   "DB_SDC_EMS_TS_1_HMI_SEK[165].EMS[1]" : UDT_SDC_EMS_TS_STAT_HMI = PLC DB_SDC_EMS_TS_1_HMI.SEK[165].EMS[1] AT %DB3810.DBX29540.0, 1 s
   "DB_SDC_EMS_TS_1_HMI_SEK[166].EMS[1]" : UDT_SDC_EMS_TS_STAT_HMI = PLC DB_SDC_EMS_TS_1_HMI.SEK[166].EMS[1] AT %DB3810.DBX29720.0, 1 s
   "DB_SDC_EMS_TS_1_HMI_SEK[167].EMS[1]" : UDT_SDC_EMS_TS_STAT_HMI = PLC DB_SDC_EMS_TS_1_HMI.SEK[167].EMS[1] AT %DB3810.DBX29900.0, 1 s
   "DB_SDC_EMS_TS_1_HMI_SEK[168].EMS[1]" : UDT_SDC_EMS_TS_STAT_HMI = PLC DB_SDC_EMS_TS_1_HMI.SEK[168].EMS[1] AT %DB3810.DBX30080.0, 1 s
   "DB_SDC_EMS_TS_1_HMI_SEK[169].EMS[1]" : UDT_SDC_EMS_TS_STAT_HMI = PLC DB_SDC_EMS_TS_1_HMI.SEK[169].EMS[1] AT %DB3810.DBX30260.0, 1 s
   "DB_SDC_EMS_TS_1_HMI_SEK[170].EMS[1]" : UDT_SDC_EMS_TS_STAT_HMI = PLC DB_SDC_EMS_TS_1_HMI.SEK[170].EMS[1] AT %DB3810.DBX30440.0, 1 s
   "DB_SDC_EMS_TS_1_HMI_SEK[190].EMS[1]" : UDT_SDC_EMS_TS_STAT_HMI = PLC DB_SDC_EMS_TS_1_HMI.SEK[190].EMS[1] AT %DB3810.DBX34040.0, 1 s
   "DB_SDC_EMS_TS_1_HMI_SEK[191].EMS[1]" : UDT_SDC_EMS_TS_STAT_HMI = PLC DB_SDC_EMS_TS_1_HMI.SEK[191].EMS[1] AT %DB3810.DBX34220.0, 1 s
   "DB_SDC_EMS_TS_1_HMI_SEK[192].EMS[1]" : UDT_SDC_EMS_TS_STAT_HMI = PLC DB_SDC_EMS_TS_1_HMI.SEK[192].EMS[1] AT %DB3810.DBX34400.0, 1 s
   "DB_SDC_EMS_TS_1_HMI_SEK[193].EMS[1]" : UDT_SDC_EMS_TS_STAT_HMI = PLC DB_SDC_EMS_TS_1_HMI.SEK[193].EMS[1] AT %DB3810.DBX34580.0, 1 s
   "DB_SDC_EMS_TS_1_HMI_SEK[194].EMS[1]" : UDT_SDC_EMS_TS_STAT_HMI = PLC DB_SDC_EMS_TS_1_HMI.SEK[194].EMS[1] AT %DB3810.DBX34760.0, 1 s
   "DB_SDC_EMS_TS_1_HMI_SEK[195].EMS[1]" : UDT_SDC_EMS_TS_STAT_HMI = PLC DB_SDC_EMS_TS_1_HMI.SEK[195].EMS[1] AT %DB3810.DBX34940.0, 1 s
   "DB_SDC_EMS_TS_1_HMI_SEK[86].EMS[1]" : UDT_SDC_EMS_TS_STAT_HMI = PLC DB_SDC_EMS_TS_1_HMI.SEK[86].EMS[1] AT %DB3810.DBX15320.0, 1 s
   "DB_SDC_EMS_TS_1_HMI_SEK[87].EMS[1]" : UDT_SDC_EMS_TS_STAT_HMI = PLC DB_SDC_EMS_TS_1_HMI.SEK[87].EMS[1] AT %DB3810.DBX15500.0, 1 s
   "DB_SDC_EMS_TS_1_HMI_SEK[137].EMS[1]" : UDT_SDC_EMS_TS_STAT_HMI = PLC DB_SDC_EMS_TS_1_HMI.SEK[137].EMS[1] AT %DB3810.DBX24500.0, 1 s
   "DB_SDC_EMS_TS_1_HMI_SEK[136].EMS[1]" : UDT_SDC_EMS_TS_STAT_HMI = PLC DB_SDC_EMS_TS_1_HMI.SEK[136].EMS[1] AT %DB3810.DBX24320.0, 1 s
   "DB_SDC_EMS_TS_1_HMI_SEK[135].EMS[1]" : UDT_SDC_EMS_TS_STAT_HMI = PLC DB_SDC_EMS_TS_1_HMI.SEK[135].EMS[1] AT %DB3810.DBX24140.0, 1 s
   "DB_SDC_EMS_TS_1_HMI_SEK[134].EMS[1]" : UDT_SDC_EMS_TS_STAT_HMI = PLC DB_SDC_EMS_TS_1_HMI.SEK[134].EMS[1] AT %DB3810.DBX23960.0, 1 s

HMI tags "DB_SDC_EMS_TS_HMI_BA2"
   "DB_SDC_EMS_TS_1_HMI_SEK[99].EMS[1]" : UDT_SDC_EMS_TS_STAT_HMI = PLC DB_SDC_EMS_TS_1_HMI.SEK[99].EMS[1] AT %DB3810.DBX17660.0, 1 s
   "DB_SDC_EMS_TS_1_HMI_SEK[100].EMS[1](1)" : UDT_SDC_EMS_TS_STAT_HMI = PLC DB_SDC_EMS_TS_1_HMI.SEK[100].EMS[1] AT %DB3810.DBX17840.0, 1 s
   "DB_SDC_EMS_TS_1_HMI_SEK[101].EMS[1](1)" : UDT_SDC_EMS_TS_STAT_HMI = PLC DB_SDC_EMS_TS_1_HMI.SEK[101].EMS[1] AT %DB3810.DBX18020.0, 1 s
   "DB_SDC_EMS_TS_1_HMI_SEK[102].EMS[1](1)" : UDT_SDC_EMS_TS_STAT_HMI = PLC DB_SDC_EMS_TS_1_HMI.SEK[102].EMS[1] AT %DB3810.DBX18200.0, 1 s
   "DB_SDC_EMS_TS_1_HMI_SEK[103].EMS[1](1)" : UDT_SDC_EMS_TS_STAT_HMI = PLC DB_SDC_EMS_TS_1_HMI.SEK[103].EMS[1] AT %DB3810.DBX18380.0, 1 s
   "DB_SDC_EMS_TS_1_HMI_SEK[104].EMS[1](1)" : UDT_SDC_EMS_TS_STAT_HMI = PLC DB_SDC_EMS_TS_1_HMI.SEK[104].EMS[1] AT %DB3810.DBX18560.0, 1 s
   "DB_SDC_EMS_TS_1_HMI_SEK[105].EMS[1](1)" : UDT_SDC_EMS_TS_STAT_HMI = PLC DB_SDC_EMS_TS_1_HMI.SEK[105].EMS[1] AT %DB3810.DBX18740.0, 1 s
   "DB_SDC_EMS_TS_1_HMI_SEK[106].EMS[1](1)" : UDT_SDC_EMS_TS_STAT_HMI = PLC DB_SDC_EMS_TS_1_HMI.SEK[106].EMS[1] AT %DB3810.DBX18920.0, 1 s
   "DB_SDC_EMS_TS_1_HMI_SEK[107].EMS[1](1)" : UDT_SDC_EMS_TS_STAT_HMI = PLC DB_SDC_EMS_TS_1_HMI.SEK[107].EMS[1] AT %DB3810.DBX19100.0, 1 s
   "DB_SDC_EMS_TS_1_HMI_SEK[108].EMS[1](1)" : UDT_SDC_EMS_TS_STAT_HMI = PLC DB_SDC_EMS_TS_1_HMI.SEK[108].EMS[1] AT %DB3810.DBX19280.0, 1 s
   "DB_SDC_EMS_TS_1_HMI_SEK[109].EMS[1](1)" : UDT_SDC_EMS_TS_STAT_HMI = PLC DB_SDC_EMS_TS_1_HMI.SEK[109].EMS[1] AT %DB3810.DBX19460.0, 1 s
   "DB_SDC_EMS_TS_1_HMI_SEK[110].EMS[1](1)" : UDT_SDC_EMS_TS_STAT_HMI = PLC DB_SDC_EMS_TS_1_HMI.SEK[110].EMS[1] AT %DB3810.DBX19640.0, 1 s
   "DB_SDC_EMS_TS_1_HMI_SEK[111].EMS[1](1)" : UDT_SDC_EMS_TS_STAT_HMI = PLC DB_SDC_EMS_TS_1_HMI.SEK[111].EMS[1] AT %DB3810.DBX19820.0, 1 s
   "DB_SDC_EMS_TS_1_HMI_SEK[112].EMS[1]" : UDT_SDC_EMS_TS_STAT_HMI = PLC DB_SDC_EMS_TS_1_HMI.SEK[112].EMS[1] AT %DB3810.DBX20000.0, 1 s
   "DB_SDC_EMS_TS_1_HMI_SEK[113].EMS[1]" : UDT_SDC_EMS_TS_STAT_HMI = PLC DB_SDC_EMS_TS_1_HMI.SEK[113].EMS[1] AT %DB3810.DBX20180.0, 1 s
   "DB_SDC_EMS_TS_1_HMI_SEK[114].EMS[1]" : UDT_SDC_EMS_TS_STAT_HMI = PLC DB_SDC_EMS_TS_1_HMI.SEK[114].EMS[1] AT %DB3810.DBX20360.0, 1 s
   "DB_SDC_EMS_TS_1_HMI_SEK[99].EMS[2]" : UDT_SDC_EMS_TS_STAT_HMI = PLC DB_SDC_EMS_TS_1_HMI.SEK[99].EMS[2] AT %DB3810.DBX17690.0, 1 s
   "DB_SDC_EMS_TS_1_HMI_SEK[100].EMS[2]" : UDT_SDC_EMS_TS_STAT_HMI = PLC DB_SDC_EMS_TS_1_HMI.SEK[100].EMS[2] AT %DB3810.DBX17870.0, 1 s
   "DB_SDC_EMS_TS_1_HMI_SEK[2]" : UDT_SDC_6EMS_TS_STAT_HMI = PLC DB_SDC_EMS_TS_1_HMI.SEK[2] AT %DB3810.DBX200.0, 1 s
   "DB_SDC_EMS_TS_1_HMI_SEK[102].EMS[2]" : UDT_SDC_EMS_TS_STAT_HMI = PLC DB_SDC_EMS_TS_1_HMI.SEK[102].EMS[2] AT %DB3810.DBX18230.0, 1 s
   "DB_SDC_EMS_TS_1_HMI_SEK[103].EMS[2]" : UDT_SDC_EMS_TS_STAT_HMI = PLC DB_SDC_EMS_TS_1_HMI.SEK[103].EMS[2] AT %DB3810.DBX18410.0, 1 s
   "DB_SDC_EMS_TS_1_HMI_SEK[104].EMS[2]" : UDT_SDC_EMS_TS_STAT_HMI = PLC DB_SDC_EMS_TS_1_HMI.SEK[104].EMS[2] AT %DB3810.DBX18590.0, 1 s
   "DB_SDC_EMS_TS_1_HMI_SEK[105].EMS[2]" : UDT_SDC_EMS_TS_STAT_HMI = PLC DB_SDC_EMS_TS_1_HMI.SEK[105].EMS[2] AT %DB3810.DBX18770.0, 1 s
   "DB_SDC_EMS_TS_1_HMI_SEK[106].EMS[2]" : UDT_SDC_EMS_TS_STAT_HMI = PLC DB_SDC_EMS_TS_1_HMI.SEK[106].EMS[2] AT %DB3810.DBX18950.0, 1 s
   "DB_SDC_EMS_TS_1_HMI_SEK[107].EMS[2]" : UDT_SDC_EMS_TS_STAT_HMI = PLC DB_SDC_EMS_TS_1_HMI.SEK[107].EMS[2] AT %DB3810.DBX19130.0, 1 s
   "DB_SDC_EMS_TS_1_HMI_SEK[108].EMS[2]" : UDT_SDC_EMS_TS_STAT_HMI = PLC DB_SDC_EMS_TS_1_HMI.SEK[108].EMS[2] AT %DB3810.DBX19310.0, 1 s
   "DB_SDC_EMS_TS_1_HMI_SEK[109].EMS[2]" : UDT_SDC_EMS_TS_STAT_HMI = PLC DB_SDC_EMS_TS_1_HMI.SEK[109].EMS[2] AT %DB3810.DBX19490.0, 1 s
   "DB_SDC_EMS_TS_1_HMI_SEK[110].EMS[2]" : UDT_SDC_EMS_TS_STAT_HMI = PLC DB_SDC_EMS_TS_1_HMI.SEK[110].EMS[2] AT %DB3810.DBX19670.0, 1 s
   "DB_SDC_EMS_TS_1_HMI_SEK[111].EMS[2]" : UDT_SDC_EMS_TS_STAT_HMI = PLC DB_SDC_EMS_TS_1_HMI.SEK[111].EMS[2] AT %DB3810.DBX19850.0, 1 s
   "DB_SDC_EMS_TS_1_HMI_SEK[112].EMS[2]" : UDT_SDC_EMS_TS_STAT_HMI = PLC DB_SDC_EMS_TS_1_HMI.SEK[112].EMS[2] AT %DB3810.DBX20030.0, 1 s
   "DB_SDC_EMS_TS_1_HMI_SEK[113].EMS[2]" : UDT_SDC_EMS_TS_STAT_HMI = PLC DB_SDC_TS_PARAMETER_4.HEADER.MAX_NR_SEK AT %DB3810.DBX20210.0, 1 s
   "DB_SDC_EMS_TS_1_HMI_SEK[114].EMS[2]" : UDT_SDC_EMS_TS_STAT_HMI = PLC DB_SDC_EMS_TS_1_HMI.SEK[114].EMS[2] AT %DB3810.DBX20390.0, 1 s
   "DB_SDC_EMS_TS_2_HMI_SEK[204].EMS[1]" : UDT_SDC_EMS_TS_STAT_HMI = PLC DB_SDC_EMS_TS_2_HMI.SEK[204].EMS[1] AT %DB3811.DBX560.0, 1 s
   "DB_SDC_EMS_TS_2_HMI_SEK[204].EMS[2]" : UDT_SDC_EMS_TS_STAT_HMI = PLC DB_SDC_EMS_TS_2_HMI.SEK[204].EMS[2] AT %DB3811.DBX590.0, 1 s
   "DB_SDC_EMS_TS_2_HMI_SEK[205].EMS[1]" : UDT_SDC_EMS_TS_STAT_HMI = PLC DB_SDC_EMS_TS_2_HMI.SEK[205].EMS[1] AT %DB3811.DBX740.0, 1 s
   "DB_SDC_EMS_TS_2_HMI_SEK[205].EMS[2]" : UDT_SDC_EMS_TS_STAT_HMI = PLC DB_SDC_EMS_TS_2_HMI.SEK[205].EMS[2] AT %DB3811.DBX770.0, 1 s
   "DB_SDC_EMS_TS_2_HMI_SEK[206].EMS[1]" : UDT_SDC_EMS_TS_STAT_HMI = PLC DB_SDC_EMS_TS_2_HMI.SEK[206].EMS[1] AT %DB3811.DBX920.0, 1 s
   "DB_SDC_EMS_TS_2_HMI_SEK[206].EMS[2]" : UDT_SDC_EMS_TS_STAT_HMI = PLC DB_SDC_EMS_TS_2_HMI.SEK[206].EMS[2] AT %DB3811.DBX950.0, 1 s
   "DB_SDC_EMS_TS_2_HMI_SEK[207].EMS[1]" : UDT_SDC_EMS_TS_STAT_HMI = PLC DB_SDC_EMS_TS_2_HMI.SEK[207].EMS[1] AT %DB3811.DBX1100.0, 1 s
   "DB_SDC_EMS_TS_2_HMI_SEK[207].EMS[2]" : UDT_SDC_EMS_TS_STAT_HMI = PLC DB_SDC_EMS_TS_2_HMI.SEK[207].EMS[2] AT %DB3811.DBX1130.0, 1 s
   "DB_SDC_EMS_TS_2_HMI_SEK[208].EMS[1]" : UDT_SDC_EMS_TS_STAT_HMI = PLC DB_SDC_EMS_TS_2_HMI.SEK[208].EMS[1] AT %DB3811.DBX1280.0, 1 s
   "DB_SDC_EMS_TS_2_HMI_SEK[208].EMS[2]" : UDT_SDC_EMS_TS_STAT_HMI = PLC DB_SDC_EMS_TS_2_HMI.SEK[208].EMS[2] AT %DB3811.DBX1310.0, 1 s
   "DB_SDC_EMS_TS_2_HMI_SEK[209].EMS[1]" : UDT_SDC_EMS_TS_STAT_HMI = PLC DB_SDC_EMS_TS_2_HMI.SEK[209].EMS[1] AT %DB3811.DBX1460.0, 1 s
   "DB_SDC_EMS_TS_2_HMI_SEK[209].EMS[2]" : UDT_SDC_EMS_TS_STAT_HMI = PLC DB_SDC_EMS_TS_2_HMI.SEK[209].EMS[2] AT %DB3811.DBX1490.0, 1 s
   "DB_SDC_EMS_TS_2_HMI_SEK[210].EMS[1]" : UDT_SDC_EMS_TS_STAT_HMI = PLC DB_SDC_EMS_TS_2_HMI.SEK[210].EMS[1] AT %DB3811.DBX1640.0, 1 s
   "DB_SDC_EMS_TS_2_HMI_SEK[210].EMS[2]" : UDT_SDC_EMS_TS_STAT_HMI = PLC DB_SDC_EMS_TS_2_HMI.SEK[210].EMS[2] AT %DB3811.DBX1670.0, 1 s
   "DB_SDC_EMS_TS_2_HMI_SEK[230].EMS[1]" : UDT_SDC_EMS_TS_STAT_HMI = PLC DB_SDC_EMS_TS_2_HMI.SEK[230].EMS[1] AT %DB3811.DBX5240.0, 1 s
   "DB_SDC_EMS_TS_2_HMI_SEK[230].EMS[2]" : UDT_SDC_EMS_TS_STAT_HMI = PLC DB_SDC_EMS_TS_2_HMI.SEK[230].EMS[2] AT %DB3811.DBX5270.0, 1 s
   "DB_SDC_EMS_TS_2_HMI_SEK[231].EMS[1]" : UDT_SDC_EMS_TS_STAT_HMI = PLC DB_SDC_EMS_TS_2_HMI.SEK[231].EMS[1] AT %DB3811.DBX5420.0, 1 s
   "DB_SDC_EMS_TS_2_HMI_SEK[231].EMS[2]" : UDT_SDC_EMS_TS_STAT_HMI = PLC DB_SDC_EMS_TS_2_HMI.SEK[231].EMS[2] AT %DB3811.DBX5450.0, 1 s
   "DB_SDC_EMS_TS_2_HMI_SEK[232].EMS[1]" : UDT_SDC_EMS_TS_STAT_HMI = PLC DB_SDC_EMS_TS_2_HMI.SEK[232].EMS[1] AT %DB3811.DBX5600.0, 1 s
   "DB_SDC_EMS_TS_2_HMI_SEK[232].EMS[2]" : UDT_SDC_EMS_TS_STAT_HMI = PLC DB_SDC_EMS_TS_2_HMI.SEK[232].EMS[2] AT %DB3811.DBX5630.0, 1 s
   "DB_SDC_EMS_TS_2_HMI_SEK[233].EMS[1]" : UDT_SDC_EMS_TS_STAT_HMI = PLC DB_SDC_EMS_TS_2_HMI.SEK[233].EMS[1] AT %DB3811.DBX5780.0, 1 s
   "DB_SDC_EMS_TS_2_HMI_SEK[233].EMS[2]" : UDT_SDC_EMS_TS_STAT_HMI = PLC DB_SDC_EMS_TS_2_HMI.SEK[233].EMS[2] AT %DB3811.DBX5810.0, 1 s
   "DB_SDC_EMS_TS_2_HMI_SEK[234].EMS[1]" : UDT_SDC_EMS_TS_STAT_HMI = PLC DB_SDC_EMS_TS_2_HMI.SEK[234].EMS[1] AT %DB3811.DBX5960.0, 1 s
   "DB_SDC_EMS_TS_2_HMI_SEK[234].EMS[2]" : UDT_SDC_EMS_TS_STAT_HMI = PLC DB_SDC_EMS_TS_2_HMI.SEK[234].EMS[2] AT %DB3811.DBX5990.0, 1 s
   "DB_SDC_EMS_TS_2_HMI_SEK[235].EMS[1]" : UDT_SDC_EMS_TS_STAT_HMI = PLC DB_SDC_EMS_TS_2_HMI.SEK[235].EMS[1] AT %DB3811.DBX6140.0, 1 s
   "DB_SDC_EMS_TS_2_HMI_SEK[235].EMS[2]" : UDT_SDC_EMS_TS_STAT_HMI = PLC DB_SDC_EMS_TS_2_HMI.SEK[235].EMS[2] AT %DB3811.DBX6170.0, 1 s

HMI tags "DB_SDC_TS_PARAMETER"
   "SDC\DB_SDC_TS_PARAMETER\DB_SDC_TS_PARAMETER_X.TS[XXX].ALLG.Pos.End_1" : DInt AT %DB0.DBD0, 1 s   // mm
   "SDC\DB_SDC_TS_PARAMETER\DB_SDC_TS_PARAMETER_X.TS[XXX].PROFIL[XX].Angle" : Int AT %DB0.DBW0, 1 s   // Setpoint: hoist position (mm)
   "DB_SDC_TS_PARAMETER_3_HEADER.DB_NR" : Int = PLC DB_SDC_TS_PARAMETER_3.HEADER.DB_NR AT %DB3706.DBW0, 1 s   // DB Nummer
   "SDC\DB_SDC_TS_PARAMETER\_TS_Par_HMI_Byte_08" : DInt, internal
   "SDC\DB_SDC_TS_PARAMETER\_TS_Par_Profil_Byte_08" : DInt, internal
   "DB_SDC_TS_PARAMETER_HMI_HEADER.LAENGE_PROFIL_DATA" : Int = PLC DB_SDC_TS_PARAMETER_HMI.HEADER.LAENGE_PROFIL_DATA AT %DB3804.DBW14, 1 s   // Länge SEK Data
   "SDC\DB_SDC_TS_PARAMETER\DB_SDC_TS_PARAMETER_X.TS[XXX].ALLG.Drive_speed_1" : DInt AT %DB0.DBD0, 1 s   // set value: drive speed (mm/min)
   "SDC\DB_SDC_TS_PARAMETER\_TS_Par_HMI_Byte_00" : DInt, internal
   "SDC\DB_SDC_TS_PARAMETER\_TS_Par_Allg_Byte_32" : DInt, internal
   "DB_SDC_TS_PARAMETER_HMI_HEADER.OFFEST_HMI_DATA" : Int = PLC DB_SDC_TS_PARAMETER_HMI.HEADER.OFFEST_HMI_DATA AT %DB3804.DBW18, 1 s   // Offestadresse der HMI SEK Data
   "SDC\DB_SDC_TS_PARAMETER\DB_SDC_TS_PARAMETER_X.TS[XXX].ALLG.Drive_speed_2" : DInt AT %DB0.DBD0, 1 s   // set value: drive speed (mm/min)
   "SDC\DB_SDC_TS_PARAMETER\DB_SDC_TS_PARAMETER_X.TS[XXX].PROFIL[XX].Tilt_offset_2" : Int AT %DB0.DBW0, 1 s   // set value: hoist offset (mm)
   "DB_SDC_TS_PARAMETER_5_HEADER.MIN_NR_SEK" : Int = PLC DB_SDC_TS_PARAMETER_5.HEADER.MIN_NR_SEK AT %DB3708.DBW2, 1 s   // Niedrigste SEK Nummer im DB
   "SDC\DB_SDC_TS_PARAMETER\DB_SDC_TS_PARAMETER_X.TS[XXX].ALLG.Stop_Position" : Int AT %DB0.DBW0, 1 s   // Stopp position, offset from start pos.(mm)
   "DB_SDC_TS_PARAMETER_HMI_HEADER.START_DAT" : Int = PLC DB_SDC_TS_PARAMETER_HMI.HEADER.START_DAT AT %DB3804.DBW6, 1 s   // Startadresse der SEK im DB
   "SDC\DB_SDC_TS_PARAMETER\_TS_Par_Allg_Byte_36" : DInt, internal
   "SDC\DB_SDC_TS_PARAMETER\_TS_Par_Allg_Byte_00" : DInt, internal
   "DB_SDC_TS_PARAMETER_5_HEADER.MAX_NR_SEK" : Int = PLC DB_SDC_TS_PARAMETER_5.HEADER.MAX_NR_SEK AT %DB3708.DBW4, 1 s   // Höchste SEK Nummer im DB
   "SDC\DB_SDC_TS_PARAMETER\_TS_Profil_Nr" : Int, internal
      on ChangeValue: "SDC_TS_PARAMETER"(); "SDC_GLOBAL_REFERENCE_PROFIL"("SDC\DB_SDC_TS_PARAMETER\_TS_Profil_Nr")
   "DB_SDC_TS_PARAMETER_HMI_HEADER.LAENGE_SEK_DATA" : Int = PLC DB_SDC_TS_PARAMETER_HMI.HEADER.LAENGE_SEK_DATA AT %DB3804.DBW8, 1 s   // Länge SEK Data
   "SDC\DB_SDC_TS_PARAMETER\DB_SDC_TS_PARAMETER_X.TS[XXX].PROFIL[XX].Tilt_offset_1" : Int AT %DB0.DBW0, 1 s   // set value: hoist offset (mm)
   "SDC\DB_SDC_TS_PARAMETER\_TS_Par_Profil_Byte_18" : DInt, internal
   "SDC\DB_SDC_TS_PARAMETER\DB_SDC_TS_PARAMETER_HMI.HMI[XX].PULT_Nr_EDIT" : Int AT %DB0.DBW0, 1 s   // Pult Nr Editieren Aktiv (HMI 1 = Master)
   "SDC\DB_SDC_TS_PARAMETER\_TS_Par_HMI_Byte_06" : DInt, internal
   "DB_SDC_TS_PARAMETER_6_HEADER.MAX_NR_SEK" : Int = PLC DB_SDC_TS_PARAMETER_6.HEADER.MAX_NR_SEK AT %DB3709.DBW4, 1 s   // Höchste SEK Nummer im DB
   "SDC\DB_SDC_TS_PARAMETER\_TS_Par_HMI_Byte_09" : DInt, internal
   "SDC\DB_SDC_TS_PARAMETER\_TS_Par_Allg_Byte_22" : DInt, internal
   "SDC\DB_SDC_TS_PARAMETER\_TS_Par_Allg_Byte_24" : DInt, internal
   "DB_SDC_TS_PARAMETER_1_HEADER.ANZ_PROFIL" : Int = PLC DB_SDC_TS_PARAMETER_1.HEADER.ANZ_PROFIL AT %DB3704.DBW10, 1 s   // Number of Profiles
   "SDC\DB_SDC_TS_PARAMETER\_TS_Par_Profil_Byte_14" : DInt, internal
   "SDC\DB_SDC_TS_PARAMETER\DB_SDC_TS_PARAMETER_HMI.HMI[XX].BILD_Nr" : Int AT %DB0.DBW0, 1 s   // Bild_Nr aktiv
   "DB_SDC_TS_PARAMETER_1_HEADER.DB_NR" : Int = PLC DB_SDC_TS_PARAMETER_1.HEADER.DB_NR AT %DB3704.DBW0, 1 s   // DB Nummer
   "SDC\DB_SDC_TS_PARAMETER\_TS_Par_Allg_Byte_27" : DInt, internal
   "DB_SDC_TS_PARAMETER_2_HEADER.MIN_NR_SEK" : Int = PLC DB_SDC_TS_PARAMETER_2.HEADER.MIN_NR_SEK AT %DB3705.DBW2, 1 s   // Niedrigste SEK Nummer im DB
   "SDC\DB_SDC_TS_PARAMETER\DB_SDC_TS_PARAMETER_X.TS[XXX].PROFIL[XX].Hoist_speed" : Int AT %DB0.DBW0, 1 s   // Setpoint: hoist speed (mm/min)
   "SDC\DB_SDC_TS_PARAMETER\_TS_Par_Allg_Byte_28" : DInt, internal
   "SDC\DB_SDC_TS_PARAMETER\_TS_Par_Profil_Byte_24" : DInt, internal
   "DB_SDC_TS_PARAMETER_1_HEADER.MAX_NR_SEK" : Int = PLC DB_SDC_TS_PARAMETER_1.HEADER.MAX_NR_SEK AT %DB3704.DBW4, 1 s   // Höchste SEK Nummer im DB
   "SDC\DB_SDC_TS_PARAMETER\_TS_Par_Allg_Byte_10" : DInt, internal
   "SDC\DB_SDC_TS_PARAMETER\_TS_Par_Profil_Byte_28" : DInt, internal
   "SDC\DB_SDC_TS_PARAMETER\DB_SDC_TS_PARAMETER_X.TS[XXX].PROFIL[XX].Tilt_Start_offset_1" : Int AT %DB0.DBW0, 1 s   // Start der Hubbewegung zu offset 1, Offset von Startpos. (mm)
   "SDC\DB_SDC_TS_PARAMETER\_TS_Par_Profil_Byte_32" : DInt, internal
   "SDC\DB_SDC_TS_PARAMETER\_TS_Par_HMI_Byte_14" : DInt, internal
   "SDC\DB_SDC_TS_PARAMETER\_TS_Par_HMI_Byte_18" : DInt, internal
   "DB_SDC_TS_PARAMETER_4_HEADER.DB_NR" : Int = PLC DB_SDC_TS_PARAMETER_4.HEADER.DB_NR AT %DB3707.DBW0, 1 s   // DB Nummer
   "DB_SDC_TS_PARAMETER_2_HEADER.DB_NR" : Int = PLC DB_SDC_TS_PARAMETER_2.HEADER.DB_NR AT %DB3705.DBW0, 1 s   // DB Nummer
   "SDC\DB_SDC_TS_PARAMETER\DB_SDC_TS_PARAMETER_X.TS[XXX].PROFIL[XX].Tilt_offset_3" : Int AT %DB0.DBW0, 1 s   // set value: hoist offset (mm)
   "SDC\DB_SDC_TS_PARAMETER\DB_SDC_TS_PARAMETER_HMI.HMI[XX].BILD_Nr_Alt" : Int AT %DB0.DBW0, 1 s   // Bild_Nr alt
   "SDC\DB_SDC_TS_PARAMETER\DB_SDC_TS_PARAMETER_HMI.HMI[XX].F_DATA" : Bool AT %DB0.DBX0.1, 1 s   // Daten Fehlerhaft
   "SDC\DB_SDC_TS_PARAMETER\DB_SDC_TS_PARAMETER_X.TS[XXX].PROFIL[XX].Tilt_offset_4" : Int AT %DB0.DBW0, 1 s   // set value: hoist offset (mm)
   "SDC\DB_SDC_TS_PARAMETER\DB_SDC_TS_PARAMETER_X.TS[XXX].PROFIL[XX].Tilt_Pos_start" : Int AT %DB0.DBW0, 1 s   // Start of hoist positioning; offset from start pos.(mm)
   "SDC\DB_SDC_TS_PARAMETER\DB_SDC_TS_PARAMETER_X.TS[XXX].ALLG.Pos.Actionpoint_1" : Int AT %DB0.DBW0, 1 s   // Antrieb Aktionspunktverschiebung1 / Drive Actionpointoffset 1
   "SDC\DB_SDC_TS_PARAMETER\_TS_Par_Allg_Byte_02" : DInt, internal
   "SDC\DB_SDC_TS_PARAMETER\DB_SDC_TS_PARAMETER_HMI.HMI[XX].PROFIL_Nr" : Int AT %DB0.DBW0, 1 s   // Profilnummer
   "SDC\DB_SDC_TS_PARAMETER\DB_SDC_TS_PARAMETER_X.TS[XXX].ALLG.Flags" : Word AT %DB0.DBW0, 1 s   // synchronous conveyor area
   "SDC\DB_SDC_TS_PARAMETER\_TS_Par_Profil_Byte_00" : DInt, internal
   "SDC\DB_SDC_TS_PARAMETER\_TS_Par_Profil_Byte_34" : DInt, internal
   "SDC\DB_SDC_TS_PARAMETER\_TS_Par_Profil_Byte_02" : DInt, internal
   "SDC\DB_SDC_TS_PARAMETER\_TS_Par_HMI_Byte_10" : DInt, internal
   "SDC\DB_SDC_TS_PARAMETER\DB_SDC_TS_PARAMETER_X.TS[XXX].PROFIL[XX].Hoist_offset_2" : Int AT %DB0.DBW0, 1 s   // set value: hoist offset (mm)
   "SDC\DB_SDC_TS_PARAMETER\_TS_Par_Profil_Byte_06" : DInt, internal
   "DB_SDC_TS_PARAMETER_4_HEADER.MAX_NR_SEK" : Int = PLC DB_SDC_TS_PARAMETER_4.HEADER.MAX_NR_SEK AT %DB3707.DBW4, 1 s   // Höchste SEK Nummer im DB
   "DB_SDC_TS_PARAMETER_HMI_HMI[1].PULT_Nr_EDIT" : Int = PLC DB_SDC_TS_PARAMETER_HMI.HMI[1].PULT_Nr_EDIT AT %DB3804.DBW20, 1 s   // Pult Nr Editieren Aktiv (HMI 1 = Master)
   "SDC\DB_SDC_TS_PARAMETER\_TS_Par_Profil_Byte_22" : DInt, internal
   "SDC\DB_SDC_TS_PARAMETER\_TS_Par_Profil_Byte_30" : DInt, internal
   "SDC\DB_SDC_TS_PARAMETER\_TS_Par_Profil_Byte_36" : DInt, internal
   "SDC\DB_SDC_TS_PARAMETER\_TS_Par_HMI_Byte_04" : DInt, internal
   "SDC\DB_SDC_TS_PARAMETER\_TS_Par_Allg_Byte_30" : DInt, internal
   "DB_SDC_TS_PARAMETER_3_HEADER.MAX_NR_SEK" : Int = PLC DB_SDC_TS_PARAMETER_3.HEADER.MAX_NR_SEK AT %DB3706.DBW4, 1 s   // Höchste SEK Nummer im DB
   "SDC\DB_SDC_TS_PARAMETER\_TS_Par_Profil_Byte_38" : DInt, internal
   "SDC\DB_SDC_TS_PARAMETER\DB_SDC_TS_PARAMETER_HMI.HMI[XX].FR_EDIT" : Bool AT %DB0.DBX0.0, 1 s   // Freigabe Editieren
   "SDC\DB_SDC_TS_PARAMETER\DB_SDC_TS_PARAMETER_X.TS[XXX].ALLG.Pos.Actionpoint_2" : Int AT %DB0.DBW0, 1 s   // Antrieb Aktionspunktverschiebung2 / Drive Actionpointoffset 2
   "SDC\DB_SDC_TS_PARAMETER\DB_SDC_TS_PARAMETER_X.TS[XXX].PROFIL[XX].Tilt_speed" : Int AT %DB0.DBW0, 1 s   // Setpoint: hoist speed (mm/min)
   "SDC\DB_SDC_TS_PARAMETER\DB_SDC_TS_PARAMETER_X.TS[XXX].PROFIL[XX].Hoist_Start_offset_3" : Int AT %DB0.DBW0, 1 s   // Start der Hubbewegung zu offset 1, Offset von Startpos. (mm)
   "SDC\DB_SDC_TS_PARAMETER\DB_SDC_TS_PARAMETER_HMI.HMI[XX].T_SAVE" : Bool AT %DB0.DBX0.2, 1 s   // Taster speichern
   "SDC\DB_SDC_TS_PARAMETER\DB_SDC_TS_PARAMETER_X.TS[XXX].ALLG.Pos.Start_1" : DInt AT %DB0.DBD0, 1 s   // mm
   "SDC\DB_SDC_TS_PARAMETER\DB_SDC_TS_PARAMETER_X.TS[XXX].PROFIL[XX].Hoist_Pos_start" : Int AT %DB0.DBW0, 1 s   // Start of hoist positioning; offset from start pos.(mm)
   "DB_SDC_TS_PARAMETER_6_HEADER.MIN_NR_SEK" : Int = PLC DB_SDC_TS_PARAMETER_6.HEADER.MIN_NR_SEK AT %DB3709.DBW2, 1 s   // Niedrigste SEK Nummer im DB
   "SDC\DB_SDC_TS_PARAMETER\_TS_Par_Allg_Byte_29" : DInt, internal
   "SDC\DB_SDC_TS_PARAMETER\DB_SDC_TS_PARAMETER_HMI.HMI[XX].SEK_Nr" : Int AT %DB0.DBW0, 1 s   // Sektionsnummer
   "SDC\DB_SDC_TS_PARAMETER\_TS_Par_Allg_Byte_26" : DInt, internal
   "SDC\DB_SDC_TS_PARAMETER\_TS_Par_Profil_Byte_42" : DInt, internal
   "SDC\DB_SDC_TS_PARAMETER\_TS_Par_Profil_Byte_20" : DInt, internal
   "SDC\DB_SDC_TS_PARAMETER\DB_SDC_TS_PARAMETER_HMI.HMI[XX].T_LOAD" : Bool AT %DB0.DBX0.3, 1 s   // Taster laden
   "DB_SDC_TS_PARAMETER_2_HEADER.MAX_NR_SEK" : Int = PLC DB_SDC_TS_PARAMETER_2.HEADER.MAX_NR_SEK AT %DB3705.DBW4, 1 s   // Höchste SEK Nummer im DB
   "SDC\DB_SDC_TS_PARAMETER\DB_SDC_TS_PARAMETER_X.TS[XXX].PROFIL[XX].Tilt_Start_offset_4" : Int AT %DB0.DBW0, 1 s   // Start der Hubbewegung zu offset 1, Offset von Startpos. (mm)
   "SDC\DB_SDC_TS_PARAMETER\_TS_Par_Profil_Byte_16" : DInt, internal
   "SDC\DB_SDC_TS_PARAMETER\DB_SDC_TS_PARAMETER_X.TS[XXX].PROFIL[XX].Tilt_Start_offset_3" : Int AT %DB0.DBW0, 1 s   // Start der Hubbewegung zu offset 1, Offset von Startpos. (mm)
   "DB_SDC_TS_PARAMETER_6_HEADER.DB_NR" : Int = PLC DB_SDC_TS_PARAMETER_6.HEADER.DB_NR AT %DB3709.DBW0, 1 s   // DB Nummer
   "SDC\DB_SDC_TS_PARAMETER\DB_SDC_TS_PARAMETER_X.TS[XXX].ALLG.Flags.DIST_VAL" : Word AT %DB0.DBW0, 1 s   // Abstandswerte / distance values
   "SDC\DB_SDC_TS_PARAMETER\DB_SDC_TS_PARAMETER_X.TS[XXX].PROFIL[XX].Tilt_Start_offset_2" : Int AT %DB0.DBW0, 1 s   // Start der Hubbewegung zu offset 1, Offset von Startpos. (mm)
   "SDC\DB_SDC_TS_PARAMETER\_TS_Par_Profil_Byte_40" : DInt, internal
   "SDC\DB_SDC_TS_PARAMETER\DB_SDC_TS_PARAMETER_X.TS[XXX].PROFIL[XX].Hoist_offset_4" : Int AT %DB0.DBW0, 1 s   // set value: hoist offset (mm)
   "SDC\DB_SDC_TS_PARAMETER\_TS_Par_HMI_Byte_12" : DInt, internal
   "SDC\DB_SDC_TS_PARAMETER\_TS_Par_Profil_Byte_12" : DInt, internal
   "SDC\DB_SDC_TS_PARAMETER\DB_SDC_TS_PARAMETER_X.TS[XXX].PROFIL[XX].Hoist_Start_offset_4" : Int AT %DB0.DBW0, 1 s   // Start der Hubbewegung zu offset 1, Offset von Startpos. (mm)
   "SDC\DB_SDC_TS_PARAMETER\_TS_Par_Profil_Byte_26" : DInt, internal
   "SDC\DB_SDC_TS_PARAMETER\DB_SDC_TS_PARAMETER_X.TS[XXX].PROFIL[XX].Hoist_Start_offset_2" : Int AT %DB0.DBW0, 1 s   // Start der Hubbewegung zu offset 1, Offset von Startpos. (mm)
   "SDC\DB_SDC_TS_PARAMETER\DB_SDC_TS_PARAMETER_X.TS[XXX].PROFIL[XX].Height" : Int AT %DB0.DBW0, 1 s   // Setpoint: hoist position (mm)
   "SDC\DB_SDC_TS_PARAMETER\_TS_DB_Nr" : Int, internal
   "SDC\DB_SDC_TS_PARAMETER\_EDIT" : Int, internal
   "SDC\DB_SDC_TS_PARAMETER\DB_SDC_TS_PARAMETER_X.TS[XXX].PROFIL[XX].Hoist_offset_3" : Int AT %DB0.DBW0, 1 s   // set value: hoist offset (mm)
   "DB_SDC_TS_PARAMETER_5_HEADER.DB_NR" : Int = PLC DB_SDC_TS_PARAMETER_5.HEADER.DB_NR AT %DB3708.DBW0, 1 s   // DB Nummer
   "SDC\DB_SDC_TS_PARAMETER\DB_SDC_TS_PARAMETER_X.TS[XXX].PROFIL[XX].Hoist_offset_1" : Int AT %DB0.DBW0, 1 s   // set value: hoist offset (mm)
   "SDC\DB_SDC_TS_PARAMETER\DB_SDC_TS_PARAMETER_HMI.HMI[XX].T_EDIT" : Bool AT %DB0.DBX0.0, 1 s   // Taster Editieren für Pult aktivieren
   "SDC\DB_SDC_TS_PARAMETER\_TS_Par_HMI_Byte_02" : DInt, internal
   "SDC\DB_SDC_TS_PARAMETER\DB_SDC_TS_PARAMETER_X.TS[XXX].PROFIL[XX].Hoist_Start_offset_1" : Int AT %DB0.DBW0, 1 s   // Start der Hubbewegung zu offset 1, Offset von Startpos. (mm)
   "SDC\DB_SDC_TS_PARAMETER\_TS_Par_Allg_Byte_06" : DInt, internal
   "DB_SDC_TS_PARAMETER_1_HEADER.MIN_NR_SEK" : Int = PLC DB_SDC_TS_PARAMETER_1.HEADER.MIN_NR_SEK AT %DB3704.DBW2, 1 s   // Niedrigste SEK Nummer im DB
   "DB_SDC_TS_PARAMETER_4_HEADER.MIN_NR_SEK" : Int = PLC DB_SDC_TS_PARAMETER_4.HEADER.MIN_NR_SEK AT %DB3707.DBW2, 1 s   // Niedrigste SEK Nummer im DB
   "DB_SDC_TS_PARAMETER_HMI_HEADER.START_HMI" : Int = PLC DB_SDC_TS_PARAMETER_HMI.HEADER.START_HMI AT %DB3804.DBW16, 1 s   // Startadresse HMI
   "DB_SDC_TS_PARAMETER_3_HEADER.MIN_NR_SEK" : Int = PLC DB_SDC_TS_PARAMETER_3.HEADER.MIN_NR_SEK AT %DB3706.DBW2, 1 s   // Niedrigste SEK Nummer im DB
   "SDC\DB_SDC_TS_PARAMETER\DB_SDC_TS_PARAMETER_HMI.HMI[XX].T_RESET_BED" : Bool AT %DB0.DBX0.1, 1 s   // Taster Reset Bedienfreigabe Pult Nr Bedienung
   "SDC\DB_SDC_TS_PARAMETER\_TS_Par_Profil_Byte_10" : DInt, internal
   "SDC\DB_SDC_TS_PARAMETER\_TS_Par_Profil_Byte_04" : DInt, internal
   "DB_SDC_TS_PARAMETER_HMI_HEADER.OFFEST_PROFIL" : Int = PLC DB_SDC_TS_PARAMETER_HMI.HEADER.OFFEST_PROFIL AT %DB3804.DBW12, 1 s   // Offestadresse der Profilparameter im TS-Parameterdatensatz
   "SDC\DB_SDC_TS_PARAMETER\DB_SDC_TS_PARAMETER_X.TS[XXX].ALLG.SEK_NEXT_1" : Int AT %DB0.DBW0, 1 s   // Sektion next 1
   "SDC\DB_SDC_TS_PARAMETER\_TS_Par_HMI_Byte_19" : DInt, internal
   "SDC\DB_SDC_TS_PARAMETER\_TS_Par_HMI_Byte_16" : DInt, internal
   "SDC\DB_SDC_TS_PARAMETER\DB_SDC_TS_PARAMETER_X.TS[XXX].ALLG.SEK_NEXT_2" : Int AT %DB0.DBW0, 1 s   // Sektion next 2
   "SDC\DB_SDC_TS_PARAMETER\_TS_Profil_Nr+1" : Int, internal
      on ChangeValue: "SDC_TS_PARAMETER"(); "SDC_GLOBAL_REFERENCE_PROFIL"("SDC\DB_SDC_TS_PARAMETER\_TS_Profil_Nr+1")
   "SDC\DB_SDC_TS_PARAMETER\DB_SDC_TS_PARAMETER_X.TS[XXX].PROFIL[XX+1].Angle" : Int AT %DB0.DBW0, 1 s   // Setpoint: hoist position (mm)
   "SDC\DB_SDC_TS_PARAMETER\DB_SDC_TS_PARAMETER_X.TS[XXX].PROFIL[XX+1].Height" : Int AT %DB0.DBW0, 1 s   // Setpoint: hoist position (mm)
   "SDC\DB_SDC_TS_PARAMETER\DB_SDC_TS_PARAMETER_X.TS[XXX].PROFIL[XX+1].Hoist_offset_1" : Int AT %DB0.DBW0, 1 s   // set value: hoist offset (mm)
   "SDC\DB_SDC_TS_PARAMETER\DB_SDC_TS_PARAMETER_X.TS[XXX].PROFIL[XX+1].Hoist_offset_2" : Int AT %DB0.DBW0, 1 s   // set value: hoist offset (mm)
   "SDC\DB_SDC_TS_PARAMETER\DB_SDC_TS_PARAMETER_X.TS[XXX].PROFIL[XX+1].Hoist_offset_3" : Int AT %DB0.DBW0, 1 s   // set value: hoist offset (mm)
   "SDC\DB_SDC_TS_PARAMETER\DB_SDC_TS_PARAMETER_X.TS[XXX].PROFIL[XX+1].Hoist_offset_4" : Int AT %DB0.DBW0, 1 s   // set value: hoist offset (mm)
   "SDC\DB_SDC_TS_PARAMETER\DB_SDC_TS_PARAMETER_X.TS[XXX].PROFIL[XX+1].Hoist_Pos_start" : Int AT %DB0.DBW0, 1 s   // Start of hoist positioning; offset from start pos.(mm)
   "SDC\DB_SDC_TS_PARAMETER\DB_SDC_TS_PARAMETER_X.TS[XXX].PROFIL[XX+1].Hoist_speed" : Int AT %DB0.DBW0, 1 s   // Setpoint: hoist speed (mm/min)
   "SDC\DB_SDC_TS_PARAMETER\DB_SDC_TS_PARAMETER_X.TS[XXX].PROFIL[XX+1].Hoist_Start_offset_1" : Int AT %DB0.DBW0, 1 s   // Start der Hubbewegung zu offset 1, Offset von Startpos. (mm)
   "SDC\DB_SDC_TS_PARAMETER\DB_SDC_TS_PARAMETER_X.TS[XXX].PROFIL[XX+1].Hoist_Start_offset_2" : Int AT %DB0.DBW0, 1 s   // Start der Hubbewegung zu offset 1, Offset von Startpos. (mm)
   "SDC\DB_SDC_TS_PARAMETER\DB_SDC_TS_PARAMETER_X.TS[XXX].PROFIL[XX+1].Hoist_Start_offset_3" : Int AT %DB0.DBW0, 1 s   // Start der Hubbewegung zu offset 1, Offset von Startpos. (mm)
   "SDC\DB_SDC_TS_PARAMETER\DB_SDC_TS_PARAMETER_X.TS[XXX].PROFIL[XX+1].Hoist_Start_offset_4" : Int AT %DB0.DBW0, 1 s   // Start der Hubbewegung zu offset 1, Offset von Startpos. (mm)
   "SDC\DB_SDC_TS_PARAMETER\DB_SDC_TS_PARAMETER_X.TS[XXX].PROFIL[XX+1].Tilt_offset_1" : Int AT %DB0.DBW0, 1 s   // set value: hoist offset (mm)
   "SDC\DB_SDC_TS_PARAMETER\DB_SDC_TS_PARAMETER_X.TS[XXX].PROFIL[XX+1].Tilt_offset_2" : Int AT %DB0.DBW0, 1 s   // set value: hoist offset (mm)
   "SDC\DB_SDC_TS_PARAMETER\DB_SDC_TS_PARAMETER_X.TS[XXX].PROFIL[XX+1].Tilt_offset_3" : Int AT %DB0.DBW0, 1 s   // set value: hoist offset (mm)
   "SDC\DB_SDC_TS_PARAMETER\DB_SDC_TS_PARAMETER_X.TS[XXX].PROFIL[XX+1].Tilt_offset_4" : Int AT %DB0.DBW0, 1 s   // set value: hoist offset (mm)
   "SDC\DB_SDC_TS_PARAMETER\DB_SDC_TS_PARAMETER_X.TS[XXX].PROFIL[XX+1].Tilt_Pos_start" : Int AT %DB0.DBW0, 1 s   // Start of hoist positioning; offset from start pos.(mm)
   "SDC\DB_SDC_TS_PARAMETER\DB_SDC_TS_PARAMETER_X.TS[XXX].PROFIL[XX+1].Tilt_speed" : Int AT %DB0.DBW0, 1 s   // Setpoint: hoist speed (mm/min)
   "SDC\DB_SDC_TS_PARAMETER\DB_SDC_TS_PARAMETER_X.TS[XXX].PROFIL[XX+1].Tilt_Start_offset_1" : Int AT %DB0.DBW0, 1 s   // Start der Hubbewegung zu offset 1, Offset von Startpos. (mm)
   "SDC\DB_SDC_TS_PARAMETER\DB_SDC_TS_PARAMETER_X.TS[XXX].PROFIL[XX+1].Tilt_Start_offset_2" : Int AT %DB0.DBW0, 1 s   // Start der Hubbewegung zu offset 1, Offset von Startpos. (mm)
   "SDC\DB_SDC_TS_PARAMETER\DB_SDC_TS_PARAMETER_X.TS[XXX].PROFIL[XX+1].Tilt_Start_offset_3" : Int AT %DB0.DBW0, 1 s   // Start der Hubbewegung zu offset 1, Offset von Startpos. (mm)
   "SDC\DB_SDC_TS_PARAMETER\DB_SDC_TS_PARAMETER_X.TS[XXX].PROFIL[XX+1].Tilt_Start_offset_4" : Int AT %DB0.DBW0, 1 s   // Start der Hubbewegung zu offset 1, Offset von Startpos. (mm)
   "SDC\DB_SDC_TS_PARAMETER\_TS_Par_Profil+1_Byte_00" : DInt, internal
   "SDC\DB_SDC_TS_PARAMETER\_TS_Par_Profil+1_Byte_02" : DInt, internal
   "SDC\DB_SDC_TS_PARAMETER\_TS_Par_Profil+1_Byte_04" : DInt, internal
   "SDC\DB_SDC_TS_PARAMETER\_TS_Par_Profil+1_Byte_06" : DInt, internal
   "SDC\DB_SDC_TS_PARAMETER\_TS_Par_Profil+1_Byte_08" : DInt, internal
   "SDC\DB_SDC_TS_PARAMETER\_TS_Par_Profil+1_Byte_10" : DInt, internal
   "SDC\DB_SDC_TS_PARAMETER\_TS_Par_Profil+1_Byte_12" : DInt, internal
   "SDC\DB_SDC_TS_PARAMETER\_TS_Par_Profil+1_Byte_14" : DInt, internal
   "SDC\DB_SDC_TS_PARAMETER\_TS_Par_Profil+1_Byte_16" : DInt, internal
   "SDC\DB_SDC_TS_PARAMETER\_TS_Par_Profil+1_Byte_18" : DInt, internal
   "SDC\DB_SDC_TS_PARAMETER\_TS_Par_Profil+1_Byte_20" : DInt, internal
   "SDC\DB_SDC_TS_PARAMETER\_TS_Par_Profil+1_Byte_22" : DInt, internal
   "SDC\DB_SDC_TS_PARAMETER\_TS_Par_Profil+1_Byte_24" : DInt, internal
   "SDC\DB_SDC_TS_PARAMETER\_TS_Par_Profil+1_Byte_26" : DInt, internal
   "SDC\DB_SDC_TS_PARAMETER\_TS_Par_Profil+1_Byte_28" : DInt, internal
   "SDC\DB_SDC_TS_PARAMETER\_TS_Par_Profil+1_Byte_30" : DInt, internal
   "SDC\DB_SDC_TS_PARAMETER\_TS_Par_Profil+1_Byte_32" : DInt, internal
   "SDC\DB_SDC_TS_PARAMETER\_TS_Par_Profil+1_Byte_34" : DInt, internal
   "SDC\DB_SDC_TS_PARAMETER\_TS_Par_Profil+1_Byte_36" : DInt, internal
   "SDC\DB_SDC_TS_PARAMETER\_TS_Par_Profil+1_Byte_38" : DInt, internal
   "SDC\DB_SDC_TS_PARAMETER\_TS_Par_Profil+1_Byte_40" : DInt, internal
   "SDC\DB_SDC_TS_PARAMETER\_TS_Par_Profil+1_Byte_42" : DInt, internal
   "DB_SDC_TS_PARAMETER_HMI_HEADER.DB_NR" : Int = PLC DB_SDC_TS_PARAMETER_HMI.HEADER.DB_NR AT %DB3804.DBW0, 1 s
   "SDC\DB_SDC_TS_PARAMETER\DB_SDC_TS_PARAMETER_HMI.HMI[XX].PROFIL_Nr_COPY" : Int AT %DB0.DBW0, 1 s   // Profilnummer
   "SDC\DB_SDC_TS_PARAMETER\DB_SDC_TS_PARAMETER_HMI.HMI[XX].PROFIL_Nr_DEST" : Int AT %DB0.DBW0, 1 s   // Profilnummer
   "SDC\DB_SDC_TS_PARAMETER\DB_SDC_TS_PARAMETER_HMI.HMI[XX].T_COPY" : Bool AT %DB0.DBX0.4, 1 s   // Taster Editieren für Pult aktivieren
   "SDC\DB_SDC_TS_PARAMETER\DB_SDC_TS_PARAMETER_HMI.HMI[XX].T_COPY_ALL" : Bool AT %DB0.DBX0.5, 1 s   // Taster Editieren für Pult aktivieren

